       "HMI_SN".pgCfg := 0;
   END_IF;
END_REGION

REGION Network 16: alm tmt
   #tim_alm[1].TON(IN := #"step".%X3 AND NOT #iB AND NOT #disAlm_Tmt, PT := #tim_alm[1].PT);
   IF #tim_alm[1].Q THEN #alm_tmt := TRUE; END_IF;
   IF ("RstAlm" AND #iB) OR #transit_end_confirmed THEN #alm_tmt := FALSE; END_IF;
   #_w1 := ("HMI_SN".instance_sel = #nrs) AND ("HMI_SN".tip_sel = 3);
   #_w2 := #_w1 AND "HMI_SN".CfOp[1];
   IF #_w2 THEN
       #alm_tmt := FALSE;
       #alm_release := FALSE;
       "HMI_SN".CfOp[1] := FALSE;
   END_IF;
   IF #_w2 AND #b0 THEN
       #mpp := TRUE;
       #alm_disapear := FALSE;
       "HMI_SN".CfOp[1] := FALSE;
       #transit_end_confirmed := TRUE;
   END_IF;
   IF #_w1 AND "HMI_SN".CfOp[2] THEN
       #mpp := FALSE;
       #alm_tmt := FALSE;
       #alm_release := FALSE;
   END_IF;
   #_w3 := #_w1 AND "HMI_SN".CfOp[2];
   IF #_w3 THEN
       "HMI_SN".CfOp[2] := FALSE;
       #transit_end_confirmed := TRUE;
   END_IF;
   IF NOT #"step".%X3 THEN #transit_end_confirmed := FALSE; END_IF;
END_REGION

REGION Network 17: alm release
   #tim_alm[2].TON(IN := #"step".%X3 AND NOT #iAr AND NOT #disAlmRls, PT := #tim_alm[2].PT);
   IF #tim_alm[2].Q THEN #alm_release := TRUE; END_IF;
   IF "RstAlm" AND #iAr THEN #alm_release := FALSE; END_IF;
END_REGION

REGION Network 18: cf op alarma disparitie fara tranzit
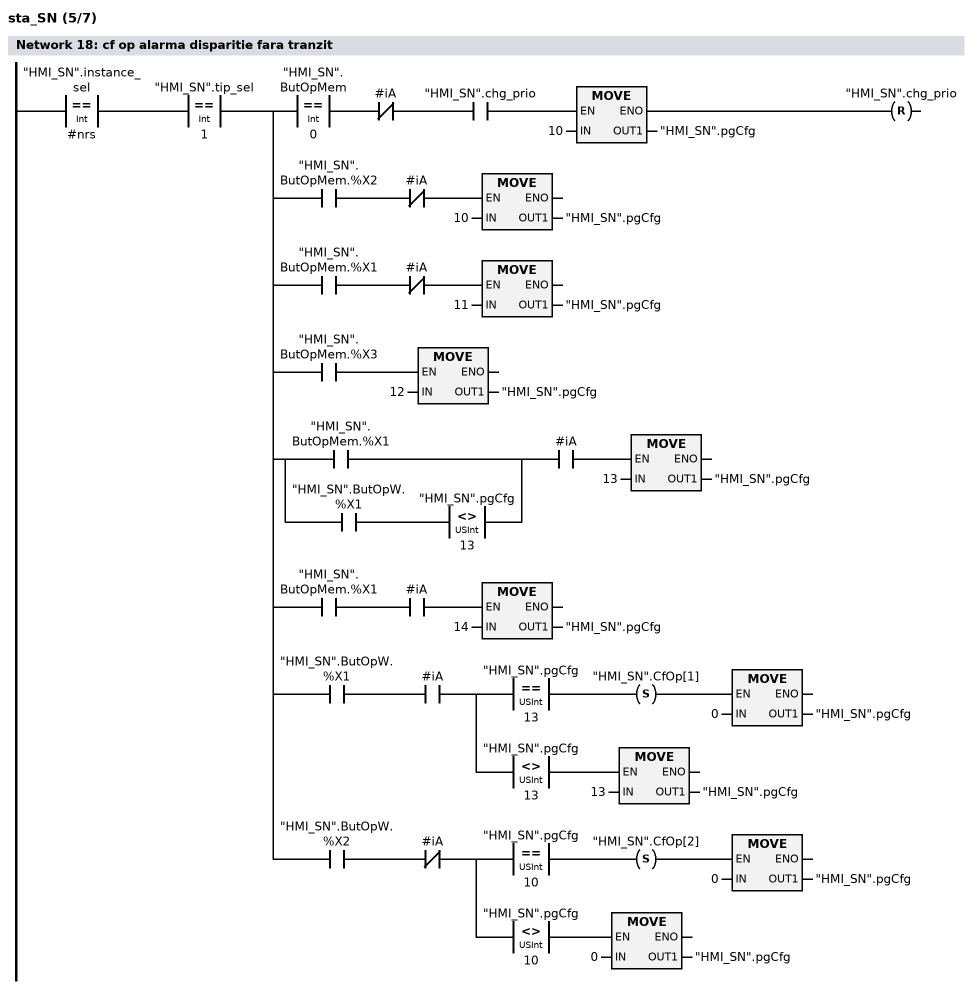
   RUNG wire#powerrail
      { S7_Templates := "SrcType := Int" } EQ_Contact(in1 := "HMI_SN".instance_sel, in2 := #nrs)
      { S7_Templates := "SrcType := Int" } EQ_Contact(in1 := "HMI_SN".tip_sel, in2 := 1)
      wire#w1
      { S7_Templates := "SrcType := Int" } EQ_Contact(in1 := "HMI_SN".ButOpMem, in2 := 0)
      I_Contact( #iA )
      Contact( "HMI_SN".chg_prio )
      Move(in := 10, out1 => "HMI_SN".pgCfg)
      R_Coil( "HMI_SN".chg_prio )
   END_RUNG
   RUNG wire#w1
      Contact( "HMI_SN".ButOpMem.%X2 )
      I_Contact( #iA )
      Move(in := 10, out1 => "HMI_SN".pgCfg)
   END_RUNG
   RUNG wire#w1
      Contact( "HMI_SN".ButOpMem.%X1 )
      I_Contact( #iA )
      Move(in := 11, out1 => "HMI_SN".pgCfg)
   END_RUNG
   RUNG wire#w1
      Contact( "HMI_SN".ButOpMem.%X3 )
      Move(in := 12, out1 => "HMI_SN".pgCfg)
   END_RUNG
   RUNG wire#w1
      Contact( "HMI_SN".ButOpMem.%X1 )
      wire#w2
      Contact( #iA )
      Move(in := 13, out1 => "HMI_SN".pgCfg)
   END_RUNG
   RUNG wire#w1
      Contact( "HMI_SN".ButOpW.%X1 )
      { S7_Templates := "SrcType := USInt" } NE_Contact(in1 := "HMI_SN".pgCfg, in2 := 13)
   END_RUNG wire#w2
   RUNG wire#w1
      Contact( "HMI_SN".ButOpMem.%X1 )
      Contact( #iA )
      Move(in := 14, out1 => "HMI_SN".pgCfg)
   END_RUNG
   RUNG wire#w1
      Contact( "HMI_SN".ButOpW.%X1 )
      Contact( #iA )
      wire#w3
      { S7_Templates := "SrcType := USInt" } EQ_Contact(in1 := "HMI_SN".pgCfg, in2 := 13)
      S_Coil( "HMI_SN".CfOp[1] )
      Move(in := 0, out1 => "HMI_SN".pgCfg)
   END_RUNG
   RUNG wire#w3
      { S7_Templates := "SrcType := USInt" } NE_Contact(in1 := "HMI_SN".pgCfg, in2 := 13)
      Move(in := 13, out1 => "HMI_SN".pgCfg)
   END_RUNG
   RUNG wire#w1
      Contact( "HMI_SN".ButOpW.%X2 )
      I_Contact( #iA )
      wire#w4
      { S7_Templates := "SrcType := USInt" } EQ_Contact(in1 := "HMI_SN".pgCfg, in2 := 10)
      S_Coil( "HMI_SN".CfOp[2] )
      Move(in := 0, out1 => "HMI_SN".pgCfg)
   END_RUNG
   RUNG wire#w4
      { S7_Templates := "SrcType := USInt" } NE_Contact(in1 := "HMI_SN".pgCfg, in2 := 10)
      Move(in := 0, out1 => "HMI_SN".pgCfg)
   END_RUNG
   // the same network as SCL:
   #_w1 := ("HMI_SN".instance_sel = #nrs) AND ("HMI_SN".tip_sel = 1);
   IF #_w1 AND ("HMI_SN".ButOpMem = 0) AND NOT #iA AND "HMI_SN".chg_prio THEN
       "HMI_SN".pgCfg := 10;
       "HMI_SN".chg_prio := FALSE;
   END_IF;
   IF #_w1 AND "HMI_SN".ButOpMem.%X2 AND NOT #iA THEN "HMI_SN".pgCfg := 10; END_IF;
   IF #_w1 AND "HMI_SN".ButOpMem.%X1 AND NOT #iA THEN "HMI_SN".pgCfg := 11; END_IF;
   IF #_w1 AND "HMI_SN".ButOpMem.%X3 THEN "HMI_SN".pgCfg := 12; END_IF;
   IF #_w1 AND ("HMI_SN".ButOpMem.%X1 OR ("HMI_SN".ButOpW.%X1 AND ("HMI_SN".pgCfg <> 13))) AND #iA THEN
       "HMI_SN".pgCfg := 13;
   END_IF;
   IF #_w1 AND "HMI_SN".ButOpMem.%X1 AND #iA THEN "HMI_SN".pgCfg := 14; END_IF;
   #_w2 := #_w1 AND "HMI_SN".ButOpW.%X1 AND #iA;
   IF #_w2 AND ("HMI_SN".pgCfg = 13) THEN
       "HMI_SN".CfOp[1] := TRUE;
       "HMI_SN".pgCfg := 0;
   END_IF;
   IF #_w2 AND ("HMI_SN".pgCfg <> 13) THEN "HMI_SN".pgCfg := 13; END_IF;
   #_w3 := #_w1 AND "HMI_SN".ButOpW.%X2 AND NOT #iA;
   IF #_w3 AND ("HMI_SN".pgCfg = 10) THEN
       "HMI_SN".CfOp[2] := TRUE;
       "HMI_SN".pgCfg := 0;
   END_IF;
   IF #_w3 AND ("HMI_SN".pgCfg <> 10) THEN "HMI_SN".pgCfg := 0; END_IF;
END_REGION

REGION Network 19: alm disap
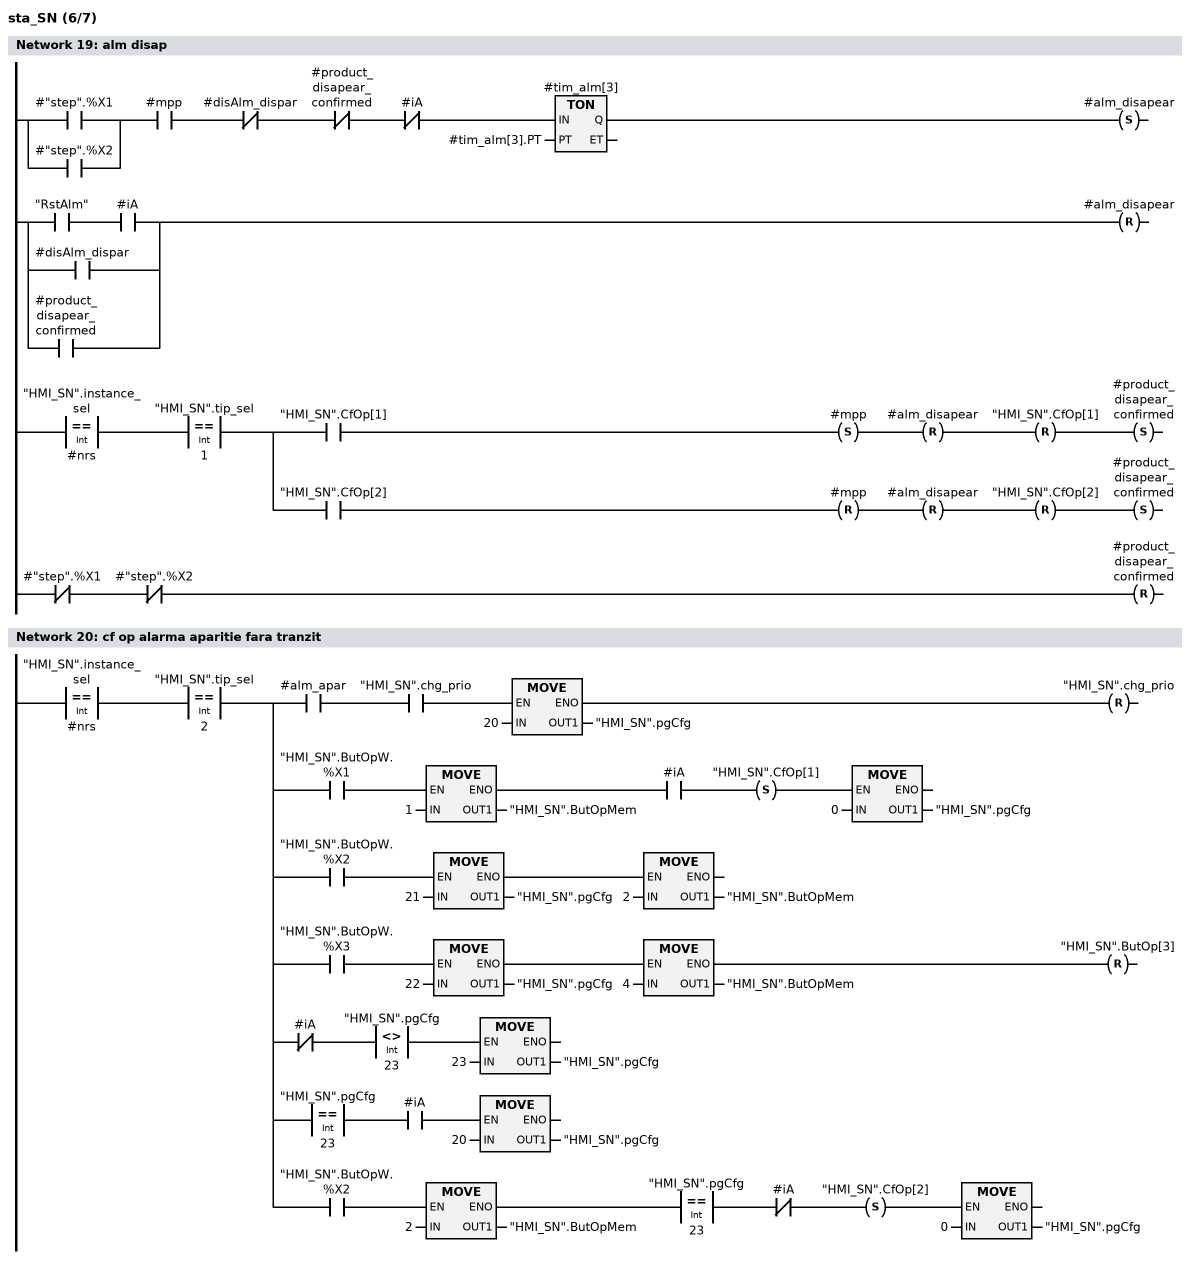
   #tim_alm[3].TON(IN := (#"step".%X1 OR #"step".%X2) AND #mpp AND NOT #disAlm_dispar AND NOT #product_disapear_confirmed AND NOT #iA,
                   PT := #tim_alm[3].PT);
   IF #tim_alm[3].Q THEN #alm_disapear := TRUE; END_IF;
   IF ("RstAlm" AND #iA) OR #disAlm_dispar OR #product_disapear_confirmed THEN
       #alm_disapear := FALSE;
   END_IF;
   #_w1 := ("HMI_SN".instance_sel = #nrs) AND ("HMI_SN".tip_sel = 1);
   IF #_w1 AND "HMI_SN".CfOp[1] THEN
       #mpp := TRUE;
       #alm_disapear := FALSE;
   END_IF;
   #_w2 := #_w1 AND "HMI_SN".CfOp[1];
   IF #_w2 THEN
       "HMI_SN".CfOp[1] := FALSE;
       #product_disapear_confirmed := TRUE;
   END_IF;
   IF #_w1 AND "HMI_SN".CfOp[2] THEN
       #mpp := FALSE;
       #alm_disapear := FALSE;
   END_IF;
   #_w3 := #_w1 AND "HMI_SN".CfOp[2];
   IF #_w3 THEN
       "HMI_SN".CfOp[2] := FALSE;
       #product_disapear_confirmed := TRUE;
   END_IF;
   IF NOT #"step".%X1 AND NOT #"step".%X2 THEN #product_disapear_confirmed := FALSE; END_IF;
END_REGION

REGION Network 20: cf op alarma aparitie fara tranzit
   RUNG wire#powerrail
      { S7_Templates := "SrcType := Int" } EQ_Contact(in1 := "HMI_SN".instance_sel, in2 := #nrs)
      { S7_Templates := "SrcType := Int" } EQ_Contact(in1 := "HMI_SN".tip_sel, in2 := 2)
      wire#w1
      Contact( #alm_apar )
      Contact( "HMI_SN".chg_prio )
      Move(in := 20, out1 => "HMI_SN".pgCfg)
      R_Coil( "HMI_SN".chg_prio )
   END_RUNG
   RUNG wire#w1
      Contact( "HMI_SN".ButOpW.%X1 )
      Move(in := 1, out1 => "HMI_SN".ButOpMem)
      Contact( #iA )
      S_Coil( "HMI_SN".CfOp[1] )
      Move(in := 0, out1 => "HMI_SN".pgCfg)
   END_RUNG
   RUNG wire#w1
      Contact( "HMI_SN".ButOpW.%X2 )
      Move(in := 21, out1 => "HMI_SN".pgCfg)
      Move(in := 2, out1 => "HMI_SN".ButOpMem)
   END_RUNG
   RUNG wire#w1
      Contact( "HMI_SN".ButOpW.%X3 )
      Move(in := 22, out1 => "HMI_SN".pgCfg)
      Move(in := 4, out1 => "HMI_SN".ButOpMem)
      R_Coil( "HMI_SN".ButOp[3] )
   END_RUNG
   RUNG wire#w1
      I_Contact( #iA )
      { S7_Templates := "SrcType := Int" } NE_Contact(in1 := "HMI_SN".pgCfg, in2 := 23)
      Move(in := 23, out1 => "HMI_SN".pgCfg)
   END_RUNG
   RUNG wire#w1
      { S7_Templates := "SrcType := Int" } EQ_Contact(in1 := "HMI_SN".pgCfg, in2 := 23)
      Contact( #iA )
      Move(in := 20, out1 => "HMI_SN".pgCfg)
   END_RUNG
   RUNG wire#w1
      Contact( "HMI_SN".ButOpW.%X2 )
      Move(in := 2, out1 => "HMI_SN".ButOpMem)
      { S7_Templates := "SrcType := Int" } EQ_Contact(in1 := "HMI_SN".pgCfg, in2 := 23)
      I_Contact( #iA )
      S_Coil( "HMI_SN".CfOp[2] )
      Move(in := 0, out1 => "HMI_SN".pgCfg)
   END_RUNG
   // the same network as SCL:
   #_w1 := ("HMI_SN".instance_sel = #nrs) AND ("HMI_SN".tip_sel = 2);
   IF #_w1 AND #alm_apar AND "HMI_SN".chg_prio THEN
       "HMI_SN".pgCfg := 20;
       "HMI_SN".chg_prio := FALSE;
   END_IF;
   #_w2 := #_w1 AND "HMI_SN".ButOpW.%X1;
   IF #_w2 THEN "HMI_SN".ButOpMem := 1; END_IF;
   IF #_w2 AND #iA THEN
       "HMI_SN".CfOp[1] := TRUE;
       "HMI_SN".pgCfg := 0;
   END_IF;
   IF #_w1 AND "HMI_SN".ButOpW.%X2 THEN
       "HMI_SN".pgCfg := 21;
       "HMI_SN".ButOpMem := 2;
   END_IF;
   IF #_w1 AND "HMI_SN".ButOpW.%X3 THEN
       "HMI_SN".pgCfg := 22;
       "HMI_SN".ButOpMem := 4;
       "HMI_SN".ButOp[3] := FALSE;
   END_IF;
   IF #_w1 AND NOT #iA AND ("HMI_SN".pgCfg <> 23) THEN "HMI_SN".pgCfg := 23; END_IF;
   IF #_w1 AND ("HMI_SN".pgCfg = 23) AND #iA THEN "HMI_SN".pgCfg := 20; END_IF;
   #_w3 := #_w1 AND "HMI_SN".ButOpW.%X2;
   IF #_w3 THEN "HMI_SN".ButOpMem := 2; END_IF;
   IF #_w3 AND ("HMI_SN".pgCfg = 23) AND NOT #iA THEN
       "HMI_SN".CfOp[2] := TRUE;
       "HMI_SN".pgCfg := 0;
   END_IF;
END_REGION

REGION Network 21: alm apar
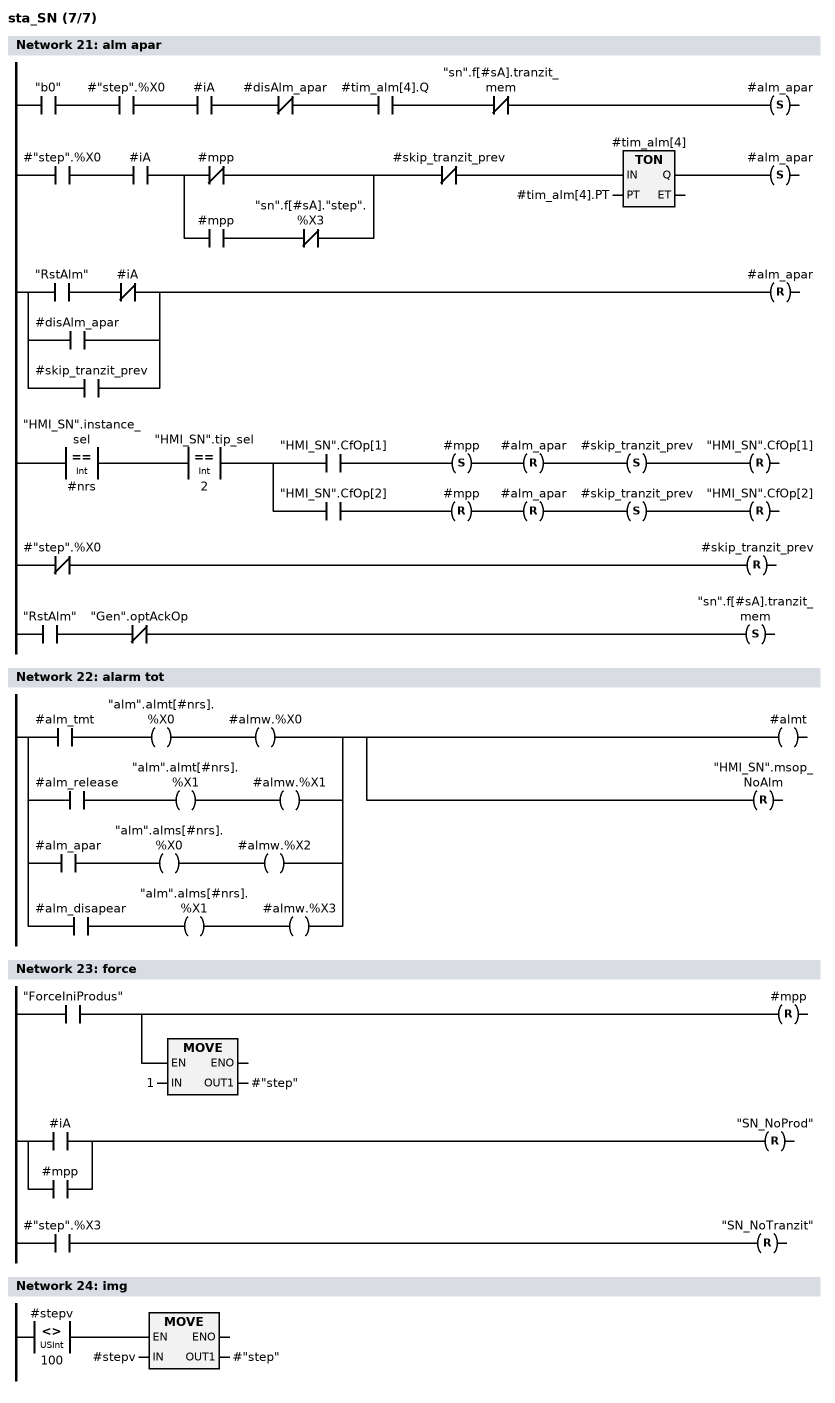
   IF "b0" AND #"step".%X0 AND #iA AND NOT #disAlm_apar AND #tim_alm[4].Q AND NOT "sn".f[#sA].tranzit_mem THEN
       #alm_apar := TRUE;
   END_IF;
   #tim_alm[4].TON(IN := #"step".%X0 AND #iA AND (NOT #mpp OR (#mpp AND NOT "sn".f[#sA]."step".%X3)) AND NOT #skip_tranzit_prev,
                   PT := #tim_alm[4].PT);
   IF #tim_alm[4].Q THEN #alm_apar := TRUE; END_IF;
   IF ("RstAlm" AND NOT #iA) OR #disAlm_apar OR #skip_tranzit_prev THEN #alm_apar := FALSE; END_IF;
   #_w1 := ("HMI_SN".instance_sel = #nrs) AND ("HMI_SN".tip_sel = 2);
   IF #_w1 AND "HMI_SN".CfOp[1] THEN
       #mpp := TRUE;
       #alm_apar := FALSE;
       #skip_tranzit_prev := TRUE;
       "HMI_SN".CfOp[1] := FALSE;
   END_IF;
   IF #_w1 AND "HMI_SN".CfOp[2] THEN
       #mpp := FALSE;
       #alm_apar := FALSE;
       #skip_tranzit_prev := TRUE;
       "HMI_SN".CfOp[2] := FALSE;
   END_IF;
   IF NOT #"step".%X0 THEN #skip_tranzit_prev := FALSE; END_IF;
   IF "RstAlm" AND NOT "Gen".optAckOp THEN "sn".f[#sA].tranzit_mem := TRUE; END_IF;
END_REGION

REGION Network 22: alarm tot
   RUNG wire#powerrail
      Contact( #alm_tmt )
      Coil( "alm".almt[#nrs].%X0 )
      Coil( #almw.%X0 )
      wire#w1
      Coil( #almt )
   END_RUNG
   RUNG wire#powerrail
      Contact( #alm_release )
      Coil( "alm".almt[#nrs].%X1 )
      Coil( #almw.%X1 )
   END_RUNG wire#w1
   RUNG wire#powerrail
      Contact( #alm_apar )
      Coil( "alm".alms[#nrs].%X0 )
      Coil( #almw.%X2 )
   END_RUNG wire#w1
   RUNG wire#powerrail
      Contact( #alm_disapear )
      Coil( "alm".alms[#nrs].%X1 )
      Coil( #almw.%X3 )
   END_RUNG wire#w1
   RUNG wire#w1
      R_Coil( "HMI_SN".msop_NoAlm )
   END_RUNG
   // the same network as SCL:
   "alm".almt[#nrs].%X0 := #alm_tmt;
   #almw.%X0 := #alm_tmt;
   "alm".almt[#nrs].%X1 := #alm_release;
   #almw.%X1 := #alm_release;
   "alm".alms[#nrs].%X0 := #alm_apar;
   #almw.%X2 := #alm_apar;
   "alm".alms[#nrs].%X1 := #alm_disapear;
   #almw.%X3 := #alm_disapear;
   #almt := #alm_tmt OR #alm_release OR #alm_apar OR #alm_disapear;
   IF #almt THEN "HMI_SN".msop_NoAlm := FALSE; END_IF;
END_REGION

REGION Network 23: force
   RUNG wire#powerrail
      Contact( "ForceIniProdus" )
      wire#w1
      R_Coil( #mpp )
   END_RUNG
   RUNG wire#w1
      Move(in := 1, out1 => #"step")
   END_RUNG
   RUNG wire#powerrail
      Contact( #iA )
      wire#w2
      R_Coil( "SN_NoProd" )
   END_RUNG
   RUNG wire#powerrail
      Contact( #mpp )
   END_RUNG wire#w2
   RUNG wire#powerrail
      Contact( #"step".%X3 )
      R_Coil( "SN_NoTranzit" )
   END_RUNG
   // the same network as SCL:
   IF "ForceIniProdus" THEN
       #mpp := FALSE;
       #"step" := 1;
   END_IF;
   IF #iA OR #mpp THEN "SN_NoProd" := FALSE; END_IF;
   IF #"step".%X3 THEN "SN_NoTranzit" := FALSE; END_IF;
END_REGION

REGION Network 24: img
   RUNG wire#powerrail
      { S7_Templates := "SrcType := USInt" } NE_Contact(in1 := #stepv, in2 := 100)
      Move(in := #stepv, out1 => #"step")
   END_RUNG
   // the same network as SCL:
   IF #stepv <> 100 THEN #"step" := #stepv; END_IF;
END_REGION
END_FUNCTION_BLOCK

// folder: log

FUNCTION "msc" : Void   // FC4, SCL
{ S7_Optimized_Access := 'TRUE' }
VERSION : 0.1
BEGIN
   IF "ms".i >= 0 AND "ms".i < "mst".sz THEN   // 0..799
       "mst".t["ms".i] := "ms".cyc *  10000 * 100 * 1000 +  "ms".tim * 100 * 1000 + "ms".v;
       "ms".vv := "mst".t["ms".i];
       "ms".i := "ms".i + 1;

   END_IF;
END_FUNCTION

FUNCTION "Main_log" : Void   // FC5, SCL
{ S7_Optimized_Access := 'TRUE' }
VERSION : 0.1
   VAR_TEMP
      d : DInt;
      dd : DInt;
      z : DInt;
   END_VAR
BEGIN
   "lad"();
   IF "ms".p100ms AND false THEN
       "ms".tv[50] := "ms".tv[50] + 1;
       IF "ms".tv[50] > 999 THEN
           "ms".tv[50] := 1;
       END_IF;
   END_IF;

   //contor timp 999.9 sec
   IF "ms".p100ms AND true THEN
       "ms".tim := "ms".tim + 1;
       IF "ms".tim > 9999 THEN
           "ms".tim := 0;
           #d := USINT_TO_DINT("FB_ProductionStatistics_DB".dat.HOUR) * 100 + "FB_ProductionStatistics_DB".dat.MINUTE;
           #z := USINT_TO_DINT("FB_ProductionStatistics_DB".dat.DAY MOD 10);
           "ms".cyc := 0;
           "ms".v :=#z * 10000 + #d ;
           "msc"();
       END_IF;
   END_IF;

   "ms".cyc := "ms".cyc + 1;
       IF "ms".cyc >=3 THEN
           "ms".cyc := 0;
       END_IF;


       "ms".tv[1].%X0 := "s".tranzit[1];
       "ms".tv[1].%X1 := "s".tranzit[2];
       "ms".tv[1].%X2 := "CS1_Start";
       "ms".tv[1].%X3 := "CS2_Start";
       "ms".tv[1].%X4 := "SCentrorMemT";
   "ms".tv[1].%X5 := 0;
   "ms".tv[1].%X6 := 0;
   "ms".tv[1].%X7 := 0;
   "ms".tv[1].%X8 := 0;

   "ms".tv[2].%X0 := "s".f[3].step.%X0;
   "ms".tv[2].%X1 := "s".f[3].step.%X1 ;
   "ms".tv[2].%X2 := "CS2_Start";
   "ms".tv[2].%X3 := "DB2_WORK_BITS".SQ_Centror_S;
   "ms".tv[2].%X4 := "s".f[3].step.%X2;
   "ms".tv[2].%X5 := "ChgLowSpd_pre";
   "ms".tv[2].%X6 := 0;
   "ms".tv[2].%X7 := 0;
   "ms".tv[2].%X8 := 0;

   "ms".tv[3].%X0 := "s".f[4].step.%X0;
   "ms".tv[3].%X1 := "ChgLowSpd";
   "ms".tv[3].%X2 := "DB2_WORK_BITS".SQ_S_Length[0];
   "ms".tv[3].%X3 := "DB2_WORK_BITS".Stacker_Handler.Input.Detectie_palet;
   "ms".tv[3].%X4 := "s".tranzit[3];
   "ms".tv[3].%X5 := "CS3_Start";
   "ms".tv[3].%X6 := "CS3_FaultAck";
   "ms".tv[3].%X7 := "s".f[4].step.%X1;
   "ms".tv[3].%X8 := "s".f[4].step.%X2;



   "ms".tv[4].%X0 := "s".tranzit[4];;
   "ms".tv[4].%X1 := "CS3_SlowSpeed";
   "ms".tv[4].%X2 := "s".f[4].step.%X3;
   "ms".tv[4].%X3 := "s".f[4].step.%X4;
       "ms".tv[4].%X4 := 0;
       "ms".tv[4].%X5 := 0;
       "ms".tv[4].%X6 := 0;
       "ms".tv[4].%X7 := 0;
       "ms".tv[4].%X8 := 0;
       //safe
       "ms".tv[5].%X0 := "DB200_SAFETY".Door_SN;
       "ms".tv[5].%X1 := "DB200_SAFETY".Door_S;
       "ms".tv[5].%X2 := "DB200_SAFETY".Mutting_Barrier_S;
       "ms".tv[5].%X3 := "DB200_SAFETY"."E-STOP_S";
       "ms".tv[5].%X4 := "DB200_SAFETY"."E-Stop_LineA";
       "ms".tv[5].%X5 := "Safe_Z2_A";
       "ms".tv[5].%X6 := "Safe_S";
       "ms".tv[5].%X7 := 0;
       "ms".tv[5].%X8 := 0;
       //energie &air
       "ms".tv[6].%X0 := "DB2_WORK_BITS".SoftStart_Zone2_A.YV1;
       "ms".tv[6].%X1 := "DB2_WORK_BITS".AG.Air;
       "ms".tv[6].%X2 := "DB2_WORK_BITS".SoftStart_Zone2_A.Sensor1 AND "DB2_WORK_BITS".SoftStart_Zone2_A.Sensor2;
       "ms".tv[6].%X3 := "DB2_WORK_BITS".SoftStart_Stacker.Sensor1 AND "DB2_WORK_BITS".SoftStart_Stacker.Sensor2;
       "ms".tv[6].%X4 := "DB2_WORK_BITS".Stacker_Drive_Handler.Input.iContactor;
       "ms".tv[6].%X5 := "DB2_WORK_BITS".Stack_Output_Drive_Handler.Input.iContactor;
       "ms".tv[6].%X6 := "Energie_S";
       "ms".tv[6].%X7 := "Energie_Z2_A";
       "ms".tv[6].%X8 := "DB_MDM_S".Energie;
       //BUT
       "ms".tv[7].%X0 := "bStart_S";
       "ms".tv[7].%X1 := "110S2";
       "ms".tv[7].%X2 := "bStop_S";
       "ms".tv[7].%X3 := "Automat_S";
       "ms".tv[7].%X4 := "RstAlm";
       "ms".tv[7].%X5 := 0;
       "ms".tv[7].%X6 := 0;
       "ms".tv[7].%X7 := 0;
       "ms".tv[7].%X8 := 0;

       "ms".tv[8].%X0 := "DB_Init_S".Init_OK;
       "ms".tv[8].%X1 := "Home_S";
       "ms".tv[8].%X2 := 0;
       "ms".tv[8].%X3 := 0;
       "ms".tv[8].%X4 := 0;
       "ms".tv[8].%X5 := 0;
       "ms".tv[8].%X6 := 0;
       "ms".tv[8].%X7 := 0;
       "ms".tv[8].%X8 := 0;
       IF false THEN



       "ms".tv[7].%X0 := 0;
       "ms".tv[7].%X1 := 0;
       "ms".tv[7].%X2 := 0;
       "ms".tv[7].%X3 := 0;
       "ms".tv[7].%X4 := 0;
       "ms".tv[7].%X5 := 0;
       "ms".tv[7].%X6 := 0;
       "ms".tv[7].%X7 := 0;
       "ms".tv[7].%X8 := 0;

       "ms".tv[8].%X0 := 0;
       "ms".tv[8].%X1 := 0;
       "ms".tv[8].%X2 := 0;
       "ms".tv[8].%X3 := 0;
       "ms".tv[8].%X4 := 0;
       "ms".tv[8].%X5 := 0;
       "ms".tv[8].%X6 := 0;
       "ms".tv[8].%X7 := 0;
       "ms".tv[8].%X8 := 0;
   END_IF;
   "ms".tv[10] := "FB_ProductionStatistics_DB".CntStack;
   "ms".tv[11] := "FB_ProductionStatistics_DB".CntPalS;
   "ms".tv[12] := "FB_ProductionStatistics_DB".CntPal;
   "ms".tv[13] := INT_TO_UINT("DB_PalletDispenser_PD2_Stacking_DB".PD1.Stepper);
   "ms".tv[14] := "DB_MDM_S".step;
   "is"();
   //"lad";
END_FUNCTION

FUNCTION "is" : Void   // FC7, SCL
{ S7_Optimized_Access := 'TRUE' }
VERSION : 0.1
   VAR_TEMP
      i : Int;
      v : DInt;
   END_VAR
BEGIN
   FOR #i := 1 TO 50 DO
       IF "ms".tv[#i] <> "ms".tvv[#i] THEN
           "ms".tvv[#i] := "ms".tv[#i];
           "ms".v := INT_TO_DINT(#i) * 1000 + "ms".tv[#i];
           "msc"();
       END_IF;
   END_FOR;
END_FUNCTION

FUNCTION "lad" : Void   // FC8, LAD
{ S7_Optimized_Access := 'TRUE' }
VERSION : 0.1
BEGIN

REGION Network 1
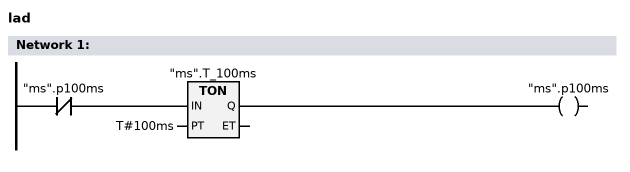
   "ms".T_100ms.TON(IN := NOT "ms".p100ms, PT := T#100ms);
   "ms".p100ms := "ms".T_100ms.Q;
END_REGION
END_FUNCTION

FUNCTION "isr" : Void   // FC9, SCL
{ S7_Optimized_Access := 'TRUE' }
VERSION : 0.1
   VAR_TEMP
      i : Int;
   END_VAR
BEGIN
   FOR #i := 0 TO 9 DO
       IF "ms".rv[#i] <> "ms".rvv[#i] THEN
           "ms".rvv[#i] := "ms".rv[#i];
           "ms".vr := INT_TO_DINT(#i) * 1000 + "ms".rv[#i];
           "mscr"();
       END_IF;
   END_FOR;
END_FUNCTION

FUNCTION "mscr" : Void   // FC10, SCL
{ S7_Optimized_Access := 'TRUE' }
VERSION : 0.1
BEGIN
   IF "ms".ir >= 0 AND "ms".ir < "mst".sz THEN   // 0..799
       "ms".rtr := USINT_TO_DINT("FB_ProductionStatistics_DB".dat.HOUR) * 100 * 100 + USINT_TO_DINT("FB_ProductionStatistics_DB".dat.MINUTE) * 100 + "FB_ProductionStatistics_DB".dat.SECOND;
    //   "mst".r["ms".ir] :="ms".rtr * 10 * 1000 + "ms".vr;
     //  "ms".vv := "mst".t["ms".i];
       "ms".ir := "ms".ir + 1;
   END_IF;
END_FUNCTION

// ===== library types =====

// folder: S7-1200/1500/Lib/S7-1200/1500/Common

FUNCTION_BLOCK "IO_LINK_DEVICE"   // FB50001, SCL
TITLE = IO_LINK_DEVICE
{ S7_Optimized_Access := 'TRUE' }
AUTHOR : SUP_FA
FAMILY : IO-Link
VERSION : 3.0
// Function block to read and write acyclic data on devices with IO-Link used on SIMATIC S7 controllers. (former IO_LINK_CALL)
   VAR_INPUT
      REQ : Bool;   // request function / Request Function / Neuer Auftrag
      ID : Hw_Io;   // hardware identifier of IO-Link master module (HW_IO) from hw-config / Hardwarekennung des IOL-Master Moduls (HW_IO) aus HW-Konfiguration
      CAP : DInt := DINT#0;   // Client Access Point (CAP), for ET200 always 227 decimal / Client Access Point (CAP), bei ET200 immer 227 dez
      RD_WR : Bool;   // read and write access on IO-Link device 0: read, 1: write / Lese und Schreibzugriff auf IO-Link Device 0: Lesen, 1: schreiben
      PORT : Int := INT#0;   // number of port on IO-Link master module (ET200SP = 0..4) / Port/ Kanalnummer an dem das IO-Link Device betrieben wird. (ET200 = 0 .. 4)
      IOL_INDEX : Int := INT#0;   // address parameter Index (IO-Link Device) 0..32767 IOL-D, 65535 port functions / Adressparameter Index (IO-Link Device) 0..32767 IOL-D, 65535 port functions
      IOL_SUBINDEX : Int := INT#0;   // address parameter Subindex (IO-Link Device) 0 full record; 1-255 single parameter / Adressparameter Subindex (IO-Link Device) 0 ges. Record; 1-255 einz. Parameter
      LEN : Int := INT#0;   // length of writing data (netto data) / Länge der zu schreibenden Daten (Nettodaten)
   END_VAR
   VAR_OUTPUT
      DONE_VALID : Bool;   // validity 0: data invalid ; 1: data valid / Gültigkeit 0: Daten nicht gültig; 1: Daten gültig
      BUSY : Bool;   // 0: request finish 1: request in progress / 0: Auftrag abgeschlossen 1: Auftrag in Bearbeitung
      ERROR : Bool;   // Error Flag = 0: no error; 1: function aborted with error / Fehler Flag 0: kein Fehler; 1: Abbruch der Funktion mit Fehler
      STATUS : DWord := DW#16#00000000;   // DP/ PNIO - error status ; ERROR Flag = 1 - communication error status in detail / DP/ PNIO - Fehlerstatus; ERROR Flag = 1 - detaillierter Kommunikationsfehlerstatus
      IOL_STATUS : DWord := DW#16#00000000;   // IO-Link error status; ERROR flag = 1: IO-Link error status in detail / IO-Link Fehlerstatus; ERROR Flag = 1 - detaillierte IO-Link Fehlerstatus
      RD_LEN : Int := INT#0;   // length of read data record (number of bytes) / Länge des gelesenen Datensatzes (Anzahl Bytes)
   END_VAR
   VAR_IN_OUT
      RECORD_IOL_DATA : Array[0..231] of Byte;   // data area for reading / writing data (max. 232 byte) / Datenbereich für LESEN / SCHREIBEN (max. 232 Byte)
   END_VAR
   VAR
      RDREC_Function : RDREC;   // system function "read data record" (former SFB52) / Funktion Datensatz lesen (ehemals SFB52)
      WRREC_Function : WRREC;   // system function "write data record" (former SFB53) / Funktion Datensatz schreiben (ehemals SFB53)
      TP_poll : TP_TIME;   // poll rate read data record / Pollzeit für "Datensatz lesen"
      TON_monitoring : TON_TIME;   // request monitoring time / Überwachungszeit für Aufträge
      rdrec : Struct   // internal structure for RDREC / interne Struktur für RDREC
         valid : Bool;   // Function performed
         busy : Bool;   // Function busy
         error : Bool;   // Error flag
         status : DWord;   // Function result/error message
         length : UInt;   // Length of the fetched data record
      END_STRUCT;
      wrrec : Struct   // internal structure for WRREC / interne Struktur für WRREC
         length : UInt;   // length of write data record
         done : Bool;   // Function performed
         busy : Bool;   // Function busy
         error : Bool;   // Error flag
         status : DWord;   // Function result/error message
      END_STRUCT;
      read : Struct   // data area for reading data / Datenbereich für Lesedaten
         header : Struct
            CALL : Struct   // header for read/write data record
               Extended_Function_Num : Byte := 16#8;   // extended function number (fix coded 08h)
               Port : Byte;   // variable port (user interface) 0...255
               FI_Index : Word := 16#FE4A;   // FI index (fix coded 65098)
            END_STRUCT;
            IOL : Struct   // header for IO-Link
               Control : Byte;   // RD_WR = 0 = read = Control:=0x03 / / RD_WR = 1 = write = Control:=0x02
               Index_HighByte : Byte;   // index of data record 0…32767 (high byte)
               Index_LowByte : Byte;   // index of data record 0…32767 (low byte)
               Subindex : Byte;   // subindex for data record 0...255
            END_STRUCT;
         END_STRUCT;
         data : Array[0..231] of Byte;
      END_STRUCT;
      write : Struct   // data area for writing data / Datenbereich für Schreibdaten
         header : Struct
            CALL : Struct   // header for read/write data record
               Extended_Function_Num : Byte := 16#8;   // extended function number (fix coded 08h)
               Port : Byte;   // variable port (user interface) 0...255
               FI_Index : Word := 16#FE4A;   // FI index (fix coded 65098)
            END_STRUCT;
            IOL : Struct   // header for IO-Link
               Control : Byte;   // RD_WR = 0 = read = Control:=0x03 / / RD_WR = 1 = write = Control:=0x02
               Index_HighByte : Byte;   // index of data record 0…32767 (high byte)
               Index_LowByte : Byte;   // index of data record 0…32767 (low byte)
               Subindex : Byte;   // subindex for data record 0...255
            END_STRUCT;
         END_STRUCT;
         data : Array[0..231] of Byte;
      END_STRUCT;
      sequencecontrol : Int := INT#0;   // number of sequence control
      typeofrequest : Int := INT#0;   // type of request (0=Read, 1=Write)
      R_TRIG_REQ : Bool;   // impulse start new request / Impuls für neuen Auftrag starten
      R_TRIG_REQ_old : Bool;   // old value of REQ (previous cycle) / Flankenmerker
      F_TRIG_poll : Bool;   // impulse poll read data record (response) / Impuls für Pollen "Datensatz lesen"
      F_TRIG_poll_old : Bool;   // old value of Poll (previous cycle) / Flankenmerker
   END_VAR
   VAR_TEMP
      retval : Int;   // function return value / Variable für Rückgabewerte von Funktionen
      tmpWORD : Word;   // data type WORD for temporarily use / Datentyp WORD zur temporären Verwendung
      tmpDWORD : DWord;   // data type DWORD for temporarily use / Datentyp DWORD zur temporären Verwendung
      tmpINT : Int;   // data type INT for temporarily use / Datentyp INT zur temporären Verwendung
      i : Int;   // run tag for counting loops / Laufvariable für for-Schleifen
   END_VAR
BEGIN
   (*---------------------------------------------------------------------------------------------------------------------
   SIEMENS AG
   ©Copyright 2015. All Rights Reserved.
   -----------------------------------------------------------------------------------------------------------------------
   Limitation of liability
   This software was developed with largest care. However, the author can not guarantee, that the software runs under
   each version of STEP7 on each PLC flawlessly.
   There is no warranty for the software, to the extent permitted by applicable law. The copyright holder provides the
   software "as is" without warranty of any kind, either expressed or implied, including, but not limited to, the implied
   warranties of merchantability and fitness for a particular purpose. The entire risk as to the quality and performance
   of the software is with you. Should the software prove defective, you assume the cost of all necessary servicing,
   repair or correction. In no event unless required by applicable law will the copyright holder be liable to you for
   damages, including any general, special, incidental or consequential damages arising out of the use or inability to
   use the software (including but not limited to loss of data or data being rendered inaccurate or losses sustained by
   you or third parties or a failure of the software to operate with any other programs), even if such holder or other
   party has been advised of the possibility of such damages.
   Permission to use or copy this software for any purpose is hereby granted without fee, provided the above notices are
   retained on all copies. Permission to modify the code and to distribute modified code is granted, provided the above
   notices are retained, and a notice that the code was modified is included with the above copyright notice.
   -----------------------------------------------------------------------------------------------------------------------
   Functionality provided by this source (short description):
   Function block IO_LINK_DEVICE - used to read and write of acyclic data records on devices with IO-Link.
   Note:
   To read data records, the IO-Link master modules needs to know which data record is required. Therefore it is necessary
   to send at first a request via write data record (only header of 8 byte). As response the IO-Link master module
   will send the required data record.

   Status:     Released (tested)
   File name:  IO_LINK_DEVICE
   System :    SIMATIC S7-1200/1500
   Version :   3.0
   -----------------------------------------------------------------------------------------------------------------------
   Script to be stored on level ... in project (mark appropriate levels with [x] below)
   [ ] External
   [ ] All levels possible
   [x] Project level
   [ ] Controller level
   [ ] Device level
   [ ] Subobject level
   -----------------------------------------------------------------------------------------------------------------------
   Restrictions, known limitations:
   The limitation of 240 byte is based on PROFIBUS DP protocol. With PROFINET IO there wouldn't no limit but because of 
   compatibility reason it wasn't changed.
     - header =   8 byte
     - data   = 232 byte
   -----------------------------------------------------------------------------------------------------------------------
   Requirements, prerequisites, External resources used: nothing
   -----------------------------------------------------------------------------------------------------------------------
   Change log table (latest change is at the bottom OF the list):
   Version Date Changes applied
   V2.0.0 <2013-09-30> First created with TIA Portal V12 SP1
   V2.1.0 <2014-03-14> Upgrade system function 'WRREC' from V1.0 to V1.1 and released for TIA Portal V13
   V3.0.0 <2015-02-28> Upgrade and released for TIA Portal V13 SP1 (without backup/restore master parameter)
   V3.0.2 <2015-07-07> Change of #IOL_INDEX and #Port lower boundry to 0
   ---------------------------------------------------------------------------------------------------------------------*)

   (*---------------------------------------------------------------------------------------------------------------------
   Description of programmed IO-Link error codes
   8000 = time out
   8001 = wrong port
   8002 = wrong index
   8003 = wrong subindex
   8005 = wrong length for write data record
   8006 = wrong length for read data record
   8052 = error during reading data record
   8053 = error during writing data record
   All other codes are coming from a higher level!
   ---------------------------------------------------------------------------------------------------------------------*)

   (*---------------------------------------------------------------------------------------------------------------------
               NEW REQUEST
   ---------------------------------------------------------------------------------------------------------------------*)
   // detection rising edge of "REQ"
   #R_TRIG_REQ := #REQ = TRUE AND #R_TRIG_REQ_old = FALSE;
   #R_TRIG_REQ_old := #REQ = TRUE;

   // start new request if not busy
   IF #R_TRIG_REQ = TRUE AND #sequencecontrol = 0 THEN
       // Freeze record ID and CAP
       #WRREC_Function.ID := #ID;
       #WRREC_Function.INDEX := #CAP;
       #RDREC_Function.ID := #ID;
       #RDREC_Function.INDEX := #CAP;

       // Initialize outputs
       #DONE_VALID := FALSE;
       #BUSY := TRUE;
       #ERROR := FALSE;
       #STATUS := DW#16#00000000;
       #IOL_STATUS := DW#16#00000000;
       #RD_LEN := INT#0;

       // Initialize data area
       #read.header.CALL.Port := B#16#0;
       #read.header.IOL.Index_LowByte := B#16#0;
       #read.header.IOL.Index_HighByte := B#16#0;
       #read.header.IOL.Subindex := B#16#0;
       #i := INT#0; // initialize loop counter      
       FOR #i := 0 TO 231 DO
           #write.data[#i] := B#16#0;
           #read.data[#i] := B#16#0;
       END_FOR;

   (*---------------------------------------------------------------------------------------------------------------------
       Setup IO-LINK Call needs a specific header
   ---------------------------------------------------------------------------------------------------------------------*)
   // setup CALL header
   #write.header.CALL.Extended_Function_Num := 16#08;  // extended function number (fix coded 08h)
   #write.header.CALL.Port := INT_TO_BYTE(#PORT);  // 1..63 = PORT number, 64..255=reserved
   #write.header.CALL.FI_Index := 65098;  // IOL-Header is following (fix coded 65098)

   // setup IOL header 
   // CONTROL = please see below at BODY
   // INDEX
   #write.header.IOL.Index_LowByte := INT_TO_BYTE(#IOL_INDEX);
   #tmpWORD := INT_TO_WORD(#IOL_INDEX);
   #tmpWORD := SHR(IN := #tmpWORD, N := 8);
   #write.header.IOL.Index_HighByte := WORD_TO_BYTE(#tmpWORD);
   // SUBINDEX
   #write.header.IOL.Subindex := INT_TO_BYTE(#IOL_SUBINDEX);